DATA_BLOCK "20_TANKS_IP_DATA"   // DB20
TITLE = Tanks Input Data
{ S7_Optimized_Access := 'TRUE' }
AUTHOR : JRS
VERSION : 0.1
// Processed data for code use
   VAR
      RIO_01 : "3T_IP_DATA";   // 1st = FPT, 2nd = 1P, 3rd = 1S
      RIO_02 : "2T_IP_DATA";   // 1st = 2P, 2nd = 2S, 3rd = N/A
      RIO_03 : "2T_IP_DATA";   // 1st = 3P, 2nd = 3S, 3rd = N/A
      RIO_04 : "2T_IP_DATA";   // BWT Level (LT-422)
      RIO_05 : "2T_IP_DATA";   // Raw minimum value from AI card
      RIO_06 : "2T_IP_DATA";   // Raw maximum value from AI card
      RIO_07 : "1T_IP_DATA";   // Normalised real value
   END_VAR
BEGIN
   RIO_02.FIRST_TANK.USD_FLOW_CNFG.ENG_MAX := 500.0;
   RIO_02.FIRST_TANK.MBG_FLOW_CNFG.ENG_MAX := 30.0;
   RIO_02.FIRST_TANK.BWT_PH_CNFG.ENG_MAX := 12.0;
   RIO_02.FIRST_TANK.O2_MONITOR_CNFG.ENG_MAX := 25.0;
   RIO_02.FIRST_TANK.DECK_IG_PRESS_CNFG.ENG_MAX := 10.0;
   RIO_02.FIRST_TANK.TANKS_PRESS_CNFG.ENG_MIN := -200.0;
   RIO_02.FIRST_TANK.TANKS_PRESS_CNFG.ENG_MAX := 200.0;
   RIO_02.FIRST_TANK.BWT_DO_CNFG.ENG_MAX := 20.0;
   RIO_02.FIRST_TANK.BWT_TEMP_CNFG.ENG_MAX := 100.0;
   RIO_02.SECOND_TANK.USD_FLOW_CNFG.ENG_MAX := 500.0;
   RIO_02.SECOND_TANK.MBG_FLOW_CNFG.ENG_MAX := 30.0;
   RIO_02.SECOND_TANK.BWT_PH_CNFG.ENG_MAX := 12.0;
   RIO_02.SECOND_TANK.BWT_DO_CNFG.ENG_MAX := 20.0;
   RIO_02.SECOND_TANK.O2_MONITOR_CNFG.ENG_MAX := 15.0;
   RIO_02.SECOND_TANK.DECK_IG_PRESS_CNFG.ENG_MAX := 25.0;
   RIO_02.SECOND_TANK.TANKS_PRESS_CNFG.ENG_MIN := -200.0;
   RIO_02.SECOND_TANK.TANKS_PRESS_CNFG.ENG_MAX := 200.0;
   RIO_02.SECOND_TANK.BWT_TEMP_CNFG.ENG_MIN := -20.0;
   RIO_02.SECOND_TANK.BWT_TEMP_CNFG.ENG_MAX := 100.0;
   RIO_02.FIRST_TANK.BWT_TEMP_CNFG.ENG_MIN := -20.0;
   RIO_02.FIRST_TANK.BWT_PH_CNFG.ENG_MIN := 2.0;
   RIO_02.SECOND_TANK.BWT_PH_CNFG.ENG_MIN := 2.0;
   RIO_01.FIRST_TANK.O2_MONITOR_CNFG.ENG_MAX := 25.0;   // Engineering units maximum value
   RIO_01.SECOND_TANK.O2_MONITOR_CNFG.ENG_MAX := 25.0;   // Engineering units maximum value
   RIO_01.THIRD_TANK.O2_MONITOR_CNFG.ENG_MAX := 25.0;   // Engineering units maximum value
   RIO_03.FIRST_TANK.O2_MONITOR_CNFG.ENG_MAX := 25.0;   // Engineering units maximum value
   RIO_03.SECOND_TANK.O2_MONITOR_CNFG.ENG_MAX := 25.0;   // Engineering units maximum value
   RIO_04.FIRST_TANK.O2_MONITOR_CNFG.ENG_MAX := 25.0;   // Engineering units maximum value
   RIO_04.SECOND_TANK.O2_MONITOR_CNFG.ENG_MAX := 25.0;   // Engineering units maximum value
   RIO_05.FIRST_TANK.O2_MONITOR_CNFG.ENG_MAX := 25.0;   // Engineering units maximum value
   RIO_05.SECOND_TANK.O2_MONITOR_CNFG.ENG_MAX := 25.0;   // Engineering units maximum value
   RIO_06.FIRST_TANK.O2_MONITOR_CNFG.ENG_MAX := 25.0;   // Engineering units maximum value
   RIO_06.SECOND_TANK.O2_MONITOR_CNFG.ENG_MAX := 25.0;   // Engineering units maximum value
   RIO_07.FIRST_TANK.O2_MONITOR_CNFG.ENG_MAX := 25.0;   // Engineering units maximum value
   RIO_07.FIRST_TANK.BWT_TEMP_CNFG.ENG_MIN := -20.0;   // Engineering units minimum value
   RIO_07.FIRST_TANK.BWT_TEMP_CNFG.ENG_MAX := 100.0;   // Engineering units maximum value
   RIO_07.FIRST_TANK.MBG_FLOW_CNFG.ENG_MAX := 30.0;   // Engineering units maximum value
   RIO_07.FIRST_TANK.USD_FLOW_CNFG.ENG_MAX := 500.0;   // Engineering units maximum value
   RIO_06.FIRST_TANK.BWT_TEMP_CNFG.ENG_MIN := -20.0;   // Engineering units minimum value
   RIO_06.FIRST_TANK.BWT_TEMP_CNFG.ENG_MAX := 100.0;   // Engineering units maximum value
   RIO_06.SECOND_TANK.BWT_TEMP_CNFG.ENG_MIN := -20.0;   // Engineering units minimum value
   RIO_06.SECOND_TANK.BWT_TEMP_CNFG.ENG_MAX := 100.0;   // Engineering units maximum value
   RIO_06.FIRST_TANK.USD_FLOW_CNFG.ENG_MAX := 500.0;   // Engineering units maximum value
   RIO_06.FIRST_TANK.MBG_FLOW_CNFG.ENG_MAX := 30.0;   // Engineering units maximum value
   RIO_06.SECOND_TANK.USD_FLOW_CNFG.ENG_MAX := 500.0;   // Engineering units maximum value
   RIO_06.SECOND_TANK.MBG_FLOW_CNFG.ENG_MAX := 30.0;   // Engineering units maximum value
   RIO_05.FIRST_TANK.BWT_TEMP_CNFG.ENG_MIN := -20.0;   // Engineering units minimum value
   RIO_05.FIRST_TANK.BWT_TEMP_CNFG.ENG_MAX := 100.0;   // Engineering units maximum value
   RIO_05.SECOND_TANK.BWT_TEMP_CNFG.ENG_MIN := -20.0;   // Engineering units minimum value
   RIO_05.SECOND_TANK.BWT_TEMP_CNFG.ENG_MAX := 100.0;   // Engineering units maximum value
   RIO_05.FIRST_TANK.USD_FLOW_CNFG.ENG_MAX := 500.0;   // Engineering units maximum value
   RIO_05.FIRST_TANK.MBG_FLOW_CNFG.ENG_MAX := 30.0;   // Engineering units maximum value
   RIO_05.SECOND_TANK.USD_FLOW_CNFG.ENG_MAX := 500.0;   // Engineering units maximum value
   RIO_05.SECOND_TANK.MBG_FLOW_CNFG.ENG_MAX := 30.0;   // Engineering units maximum value
   RIO_04.FIRST_TANK.USD_FLOW_CNFG.ENG_MAX := 500.0;   // Engineering units maximum value
   RIO_04.FIRST_TANK.MBG_FLOW_CNFG.ENG_MAX := 30.0;   // Engineering units maximum value
   RIO_04.FIRST_TANK.BWT_TEMP_CNFG.ENG_MIN := -20.0;   // Engineering units minimum value
   RIO_04.FIRST_TANK.BWT_TEMP_CNFG.ENG_MAX := 100.0;   // Engineering units maximum value
   RIO_04.SECOND_TANK.USD_FLOW_CNFG.ENG_MAX := 500.0;   // Engineering units maximum value
   RIO_04.SECOND_TANK.MBG_FLOW_CNFG.ENG_MAX := 30.0;   // Engineering units maximum value
   RIO_04.SECOND_TANK.BWT_TEMP_CNFG.ENG_MIN := -20.0;   // Engineering units minimum value
   RIO_04.SECOND_TANK.BWT_TEMP_CNFG.ENG_MAX := 100.0;   // Engineering units maximum value
   RIO_03.FIRST_TANK.USD_FLOW_CNFG.ENG_MAX := 500.0;   // Engineering units maximum value
   RIO_03.FIRST_TANK.MBG_FLOW_CNFG.ENG_MAX := 30.0;   // Engineering units maximum value
   RIO_03.FIRST_TANK.BWT_TEMP_CNFG.ENG_MIN := -20.0;   // Engineering units minimum value
   RIO_03.FIRST_TANK.BWT_TEMP_CNFG.ENG_MAX := 100.0;   // Engineering units maximum value
   RIO_01.FIRST_TANK.USD_FLOW_CNFG.ENG_MAX := 500.0;   // Engineering units maximum value
   RIO_01.FIRST_TANK.MBG_FLOW_CNFG.ENG_MAX := 30.0;   // Engineering units maximum value
   RIO_01.FIRST_TANK.BWT_TEMP_CNFG.ENG_MIN := -20.0;   // Engineering units minimum value
   RIO_01.FIRST_TANK.BWT_TEMP_CNFG.ENG_MAX := 100.0;   // Engineering units maximum value
   RIO_01.SECOND_TANK.USD_FLOW_CNFG.ENG_MAX := 500.0;   // Engineering units maximum value
   RIO_01.SECOND_TANK.MBG_FLOW_CNFG.ENG_MAX := 30.0;   // Engineering units maximum value
   RIO_01.SECOND_TANK.BWT_TEMP_CNFG.ENG_MIN := -20.0;   // Engineering units minimum value
   RIO_01.SECOND_TANK.BWT_TEMP_CNFG.ENG_MAX := 100.0;   // Engineering units maximum value
   RIO_01.THIRD_TANK.USD_FLOW_CNFG.ENG_MAX := 500.0;   // Engineering units maximum value
   RIO_01.THIRD_TANK.MBG_FLOW_CNFG.ENG_MAX := 30.0;   // Engineering units maximum value
   RIO_01.THIRD_TANK.BWT_TEMP_CNFG.ENG_MIN := -20.0;   // Engineering units minimum value
   RIO_01.THIRD_TANK.BWT_TEMP_CNFG.ENG_MAX := 100.0;   // Engineering units maximum value
   RIO_03.SECOND_TANK.USD_FLOW_CNFG.ENG_MAX := 500.0;   // Engineering units maximum value
   RIO_03.SECOND_TANK.MBG_FLOW_CNFG.ENG_MAX := 30.0;   // Engineering units maximum value
   // RIO_02.FIRST_TANK.USD_FLOW_CNFG : IW160 - USD Flow (FIT-418) - Tank #1
   // RIO_02.FIRST_TANK.MBG_FLOW_CNFG : IW162 - MBG Flow (FIT-420) - Tank #1
   // RIO_02.FIRST_TANK.BWT_LEVEL_CNFG : BWT Level (LT-422)
   // RIO_02.FIRST_TANK.BWT_PH_CNFG : BWT Ph (426)
   // RIO_02.FIRST_TANK.BWT_TEMP_CNFG : BWT Temperature (426)
   // RIO_02.FIRST_TANK.BWT_DO_CNFG : BWT DO (428)
   // RIO_02.FIRST_TANK.O2_MONITOR_CNFG : O2 Monitor (600-Tx-433)
   // RIO_02.FIRST_TANK.DECK_IG_PRESS_CNFG : Deck Main IG Pressure (PT-415)
   // RIO_02.FIRST_TANK.TANKS_PRESS_CNFG : Tank Group Pressure (PT-424)
   // RIO_02.SECOND_TANK.USD_FLOW_CNFG : IW160 - USD Flow (FIT-417) - Tank #1
   // RIO_02.SECOND_TANK.MBG_FLOW_CNFG : IW162 - MBG Flow (FIT-419) - Tank #1
   // RIO_02.SECOND_TANK.BWT_LEVEL_CNFG : BWT Level (LT-422)
   // RIO_02.SECOND_TANK.BWT_PH_CNFG : BWT Ph (426)
   // RIO_02.SECOND_TANK.BWT_TEMP_CNFG : BWT Temperature (426)
   // RIO_02.SECOND_TANK.BWT_DO_CNFG : BWT DO (428)
   // RIO_02.SECOND_TANK.SPARE_AI_1_CNFG : Input processing configuration data
   // RIO_02.SECOND_TANK.SPARE_AI_2_CNFG : Input processing configuration data
   // RIO_02.SECOND_TANK.SPARE_AI_3_CNFG : Input processing configuration data
   // RIO_02.SECOND_TANK.O2_MONITOR_CNFG : O2 Monitor (600-Tx-433)
   // RIO_02.SECOND_TANK.DECK_IG_PRESS_CNFG : Deck Main IG Pressure (PT-415)
   // RIO_02.SECOND_TANK.TANKS_PRESS_CNFG : Tank Group Pressure (PT-424)
   // RIO_02.SECOND_TANK.MBG_FLOW : FIT-419
   // RIO_02.SECOND_TANK.USD_FLOW : FIT-417
   // RIO_01.FIRST_TANK.O2_MONITOR : Space monitor, 600-Tx-433
   // RIO_01.FIRST_TANK.DECK_IG_PRESS : Deck main IG pressure, PT-415
   // RIO_01.FIRST_TANK.TANKS_PRESS : Tank group pressure, PT-424
   // RIO_01.FIRST_TANK.TANKS_PRESS_HIHI : Tank group pressure, PS-436
   // RIO_01.FIRST_TANK.TANK_GROUP_SPARE_DI_2 : Spare input
   // RIO_01.FIRST_TANK.TANK_GROUP_SPARE_DI_3 : Spare input
   // RIO_01.FIRST_TANK.TANK_GROUP_SPARE_DI_4 : Spare input
   // RIO_01.FIRST_TANK.TANK_GROUP_SPARE_DI_5 : Spare input
   // RIO_01.FIRST_TANK.TANK_GROUP_SPARE_DI_6 : Spare input
   // RIO_01.FIRST_TANK.TANK_GROUP_SPARE_DI_7 : Spare input
   // RIO_01.FIRST_TANK.GTT_ISOL_VALVE_OPEN : Gas to tank isolation valve feedback, CV-422
   // RIO_01.FIRST_TANK.GTT_ISOL_VALVE_CLSD : Gas to tank isolation valve feedback, CV-422
   // RIO_01.FIRST_TANK.TANK_VENT_A_OPEN : Tank vent valve feedback, CV-441-A
   // RIO_01.FIRST_TANK.TANK_VENT_A_CLSD : Tank vent valve feedback, CV-441-A
   // RIO_01.FIRST_TANK.TANK_VENT_B_OPEN : Tank vent valve feedback, CV-441-B
   // RIO_01.FIRST_TANK.TANK_VENT_B_CLSD : Tank vent valve feedback, CV-441-B
   // RIO_01.FIRST_TANK.BWT_LEVEL_HIHI : Tank water level, LS-425
   // RIO_01.FIRST_TANK.TANK_ALARM : Spare input
   // RIO_01.FIRST_TANK.SPARE_DI_7 : Spare input
   // RIO_01.FIRST_TANK.USD_FLOW : FIT-418
   // RIO_01.FIRST_TANK.MBG_FLOW : FIT-420
   // RIO_01.FIRST_TANK.BWT_LEVEL : LT-422
   // RIO_01.FIRST_TANK.BWT_PH : Ph 426
   // RIO_01.FIRST_TANK.BWT_TEMP : Temperature 426
   // RIO_01.FIRST_TANK.BWT_DO : Disolved oxygen 428
   // RIO_01.FIRST_TANK.SPARE_AI_1 : Spare input
   // RIO_01.FIRST_TANK.SPARE_AI_2 : Spare input
   // RIO_01.FIRST_TANK.SPARE_AI_3 : Spare input
   // RIO_01.FIRST_TANK.USD_FLOW_CNFG : IW160 - USD Flow (FIT-418) - Tank #1
   // RIO_01.FIRST_TANK.USD_FLOW_CNFG.RAW_MIN : Raw minimum value from AI card
   // RIO_01.FIRST_TANK.USD_FLOW_CNFG.RAW_MAX : Raw maximum value from AI card
   // RIO_01.FIRST_TANK.USD_FLOW_CNFG.NORM : Normalised real value
   // RIO_01.FIRST_TANK.USD_FLOW_CNFG.ENG_MIN : Engineering units minimum value
   // RIO_01.FIRST_TANK.MBG_FLOW_CNFG : IW162 - MBG Flow (FIT-420) - Tank #1
   // RIO_01.FIRST_TANK.MBG_FLOW_CNFG.RAW_MIN : Raw minimum value from AI card
   // RIO_01.FIRST_TANK.MBG_FLOW_CNFG.RAW_MAX : Raw maximum value from AI card
   // RIO_01.FIRST_TANK.MBG_FLOW_CNFG.NORM : Normalised real value
   // RIO_01.FIRST_TANK.MBG_FLOW_CNFG.ENG_MIN : Engineering units minimum value
   // RIO_01.FIRST_TANK.BWT_LEVEL_CNFG : BWT Level (LT-422)
   // RIO_01.FIRST_TANK.BWT_LEVEL_CNFG.RAW_MIN : Raw minimum value from AI card
   // RIO_01.FIRST_TANK.BWT_LEVEL_CNFG.RAW_MAX : Raw maximum value from AI card
   // RIO_01.FIRST_TANK.BWT_LEVEL_CNFG.NORM : Normalised real value
   // RIO_01.FIRST_TANK.BWT_LEVEL_CNFG.ENG_MIN : Engineering units minimum value
   // RIO_01.FIRST_TANK.BWT_LEVEL_CNFG.ENG_MAX : Engineering units maximum value
   // RIO_01.FIRST_TANK.BWT_PH_CNFG : BWT Ph (426)
   // RIO_01.FIRST_TANK.BWT_PH_CNFG.RAW_MIN : Raw minimum value from AI card
   // RIO_01.FIRST_TANK.BWT_PH_CNFG.RAW_MAX : Raw maximum value from AI card
   // RIO_01.FIRST_TANK.BWT_PH_CNFG.NORM : Normalised real value
   // RIO_01.FIRST_TANK.BWT_PH_CNFG.ENG_MIN : Engineering units minimum value
   // RIO_01.FIRST_TANK.BWT_PH_CNFG.ENG_MAX : Engineering units maximum value
   // RIO_01.FIRST_TANK.BWT_TEMP_CNFG : BWT Temperature (426)
   // RIO_01.FIRST_TANK.BWT_TEMP_CNFG.RAW_MIN : Raw minimum value from AI card
   // RIO_01.FIRST_TANK.BWT_TEMP_CNFG.RAW_MAX : Raw maximum value from AI card
   // RIO_01.FIRST_TANK.BWT_TEMP_CNFG.NORM : Normalised real value
   // RIO_01.FIRST_TANK.BWT_DO_CNFG : BWT DO (428)
   // RIO_01.FIRST_TANK.BWT_DO_CNFG.RAW_MIN : Raw minimum value from AI card
   // RIO_01.FIRST_TANK.BWT_DO_CNFG.RAW_MAX : Raw maximum value from AI card
   // RIO_01.FIRST_TANK.BWT_DO_CNFG.NORM : Normalised real value
   // RIO_01.FIRST_TANK.BWT_DO_CNFG.ENG_MIN : Engineering units minimum value
   // RIO_01.FIRST_TANK.BWT_DO_CNFG.ENG_MAX : Engineering units maximum value
   // RIO_01.FIRST_TANK.SPARE_AI_1_CNFG : Input processing configuration data
   // RIO_01.FIRST_TANK.SPARE_AI_1_CNFG.RAW_MIN : Raw minimum value from AI card
   // RIO_01.FIRST_TANK.SPARE_AI_1_CNFG.RAW_MAX : Raw maximum value from AI card
   // RIO_01.FIRST_TANK.SPARE_AI_1_CNFG.NORM : Normalised real value
   // RIO_01.FIRST_TANK.SPARE_AI_1_CNFG.ENG_MIN : Engineering units minimum value
   // RIO_01.FIRST_TANK.SPARE_AI_1_CNFG.ENG_MAX : Engineering units maximum value
   // RIO_01.FIRST_TANK.SPARE_AI_2_CNFG : Input processing configuration data
   // RIO_01.FIRST_TANK.SPARE_AI_2_CNFG.RAW_MIN : Raw minimum value from AI card
   // RIO_01.FIRST_TANK.SPARE_AI_2_CNFG.RAW_MAX : Raw maximum value from AI card
   // RIO_01.FIRST_TANK.SPARE_AI_2_CNFG.NORM : Normalised real value
   // RIO_01.FIRST_TANK.SPARE_AI_2_CNFG.ENG_MIN : Engineering units minimum value
   // RIO_01.FIRST_TANK.SPARE_AI_2_CNFG.ENG_MAX : Engineering units maximum value
   // RIO_01.FIRST_TANK.SPARE_AI_3_CNFG : Input processing configuration data
   // RIO_01.FIRST_TANK.SPARE_AI_3_CNFG.RAW_MIN : Raw minimum value from AI card
   // RIO_01.FIRST_TANK.SPARE_AI_3_CNFG.RAW_MAX : Raw maximum value from AI card
   // RIO_01.FIRST_TANK.SPARE_AI_3_CNFG.NORM : Normalised real value
   // RIO_01.FIRST_TANK.SPARE_AI_3_CNFG.ENG_MIN : Engineering units minimum value
   // RIO_01.FIRST_TANK.SPARE_AI_3_CNFG.ENG_MAX : Engineering units maximum value
   // RIO_01.FIRST_TANK.O2_MONITOR_CNFG : O2 Monitor (600-Tx-433)
   // RIO_01.FIRST_TANK.O2_MONITOR_CNFG.RAW_MIN : Raw minimum value from AI card
   // RIO_01.FIRST_TANK.O2_MONITOR_CNFG.RAW_MAX : Raw maximum value from AI card
   // RIO_01.FIRST_TANK.O2_MONITOR_CNFG.NORM : Normalised real value
   // RIO_01.FIRST_TANK.O2_MONITOR_CNFG.ENG_MIN : Engineering units minimum value
   // RIO_01.FIRST_TANK.DECK_IG_PRESS_CNFG : Deck Main IG Pressure (PT-415)
   // RIO_01.FIRST_TANK.DECK_IG_PRESS_CNFG.RAW_MIN : Raw minimum value from AI card
   // RIO_01.FIRST_TANK.DECK_IG_PRESS_CNFG.RAW_MAX : Raw maximum value from AI card
   // RIO_01.FIRST_TANK.DECK_IG_PRESS_CNFG.NORM : Normalised real value
   // RIO_01.FIRST_TANK.DECK_IG_PRESS_CNFG.ENG_MIN : Engineering units minimum value
   // RIO_01.FIRST_TANK.DECK_IG_PRESS_CNFG.ENG_MAX : Engineering units maximum value
   // RIO_01.FIRST_TANK.TANKS_PRESS_CNFG : Tank Group Pressure (PT-424)
   // RIO_01.FIRST_TANK.TANKS_PRESS_CNFG.RAW_MIN : Raw minimum value from AI card
   // RIO_01.FIRST_TANK.TANKS_PRESS_CNFG.RAW_MAX : Raw maximum value from AI card
   // RIO_01.FIRST_TANK.TANKS_PRESS_CNFG.NORM : Normalised real value
   // RIO_01.FIRST_TANK.TANKS_PRESS_CNFG.ENG_MIN : Engineering units minimum value
   // RIO_01.FIRST_TANK.TANKS_PRESS_CNFG.ENG_MAX : Engineering units maximum value
   // RIO_01.THIRD_TANK.O2_MONITOR : Space monitor, 600-Tx-433
   // RIO_01.THIRD_TANK.DECK_IG_PRESS : Deck main IG pressure, PT-415
   // RIO_01.THIRD_TANK.TANKS_PRESS : Tank group pressure, PT-424
   // RIO_01.THIRD_TANK.TANKS_PRESS_HIHI : Tank group pressure, PS-436
   // RIO_01.THIRD_TANK.TANK_GROUP_SPARE_DI_2 : Spare input
   // RIO_01.THIRD_TANK.TANK_GROUP_SPARE_DI_3 : Spare input
   // RIO_01.THIRD_TANK.TANK_GROUP_SPARE_DI_4 : Spare input
   // RIO_01.THIRD_TANK.TANK_GROUP_SPARE_DI_5 : Spare input
   // RIO_01.THIRD_TANK.TANK_GROUP_SPARE_DI_6 : Spare input
   // RIO_01.THIRD_TANK.TANK_GROUP_SPARE_DI_7 : Spare input
   // RIO_01.THIRD_TANK.GTT_ISOL_VALVE_OPEN : Gas to tank isolation valve feedback, CV-422
   // RIO_01.THIRD_TANK.GTT_ISOL_VALVE_CLSD : Gas to tank isolation valve feedback, CV-422
   // RIO_01.THIRD_TANK.TANK_VENT_A_OPEN : Tank vent valve feedback, CV-441-A
   // RIO_01.THIRD_TANK.TANK_VENT_A_CLSD : Tank vent valve feedback, CV-441-A
   // RIO_01.THIRD_TANK.TANK_VENT_B_OPEN : Tank vent valve feedback, CV-441-B
   // RIO_01.THIRD_TANK.TANK_VENT_B_CLSD : Tank vent valve feedback, CV-441-B
   // RIO_01.THIRD_TANK.BWT_LEVEL_HIHI : Tank water level, LS-425
   // RIO_01.THIRD_TANK.TANK_ALARM : Spare input
   // RIO_01.THIRD_TANK.SPARE_DI_7 : Spare input
   // RIO_01.THIRD_TANK.USD_FLOW : FIT-417
   // RIO_01.THIRD_TANK.MBG_FLOW : FIT-419
   // RIO_01.THIRD_TANK.BWT_LEVEL : LT-422
   // RIO_01.THIRD_TANK.BWT_PH : Ph 426
   // RIO_01.THIRD_TANK.BWT_TEMP : Temperature 426
   // RIO_01.THIRD_TANK.BWT_DO : Disolved oxygen 428
   // RIO_01.THIRD_TANK.SPARE_AI_1 : Spare input
   // RIO_01.THIRD_TANK.SPARE_AI_2 : Spare input
   // RIO_01.THIRD_TANK.SPARE_AI_3 : Spare input
   // RIO_01.THIRD_TANK.USD_FLOW_CNFG : IW160 - USD Flow (FIT-417) - Tank #1
   // RIO_01.THIRD_TANK.USD_FLOW_CNFG.RAW_MIN : Raw minimum value from AI card
   // RIO_01.THIRD_TANK.USD_FLOW_CNFG.RAW_MAX : Raw maximum value from AI card
   // RIO_01.THIRD_TANK.USD_FLOW_CNFG.NORM : Normalised real value
   // RIO_01.THIRD_TANK.USD_FLOW_CNFG.ENG_MIN : Engineering units minimum value
   // RIO_01.THIRD_TANK.MBG_FLOW_CNFG : IW162 - MBG Flow (FIT-420) - Tank #1
   // RIO_01.THIRD_TANK.MBG_FLOW_CNFG.RAW_MIN : Raw minimum value from AI card
   // RIO_01.THIRD_TANK.MBG_FLOW_CNFG.RAW_MAX : Raw maximum value from AI card
   // RIO_01.THIRD_TANK.MBG_FLOW_CNFG.NORM : Normalised real value
   // RIO_01.THIRD_TANK.MBG_FLOW_CNFG.ENG_MIN : Engineering units minimum value
   // RIO_01.THIRD_TANK.BWT_LEVEL_CNFG : BWT Level (LT-422)
   // RIO_01.THIRD_TANK.BWT_LEVEL_CNFG.RAW_MIN : Raw minimum value from AI card
   // RIO_01.THIRD_TANK.BWT_LEVEL_CNFG.RAW_MAX : Raw maximum value from AI card
   // RIO_01.THIRD_TANK.BWT_LEVEL_CNFG.NORM : Normalised real value
   // RIO_01.THIRD_TANK.BWT_LEVEL_CNFG.ENG_MIN : Engineering units minimum value
   // RIO_01.THIRD_TANK.BWT_LEVEL_CNFG.ENG_MAX : Engineering units maximum value
   // RIO_01.THIRD_TANK.BWT_PH_CNFG : BWT Ph (426)
   // RIO_01.THIRD_TANK.BWT_PH_CNFG.RAW_MIN : Raw minimum value from AI card
   // RIO_01.THIRD_TANK.BWT_PH_CNFG.RAW_MAX : Raw maximum value from AI card
   // RIO_01.THIRD_TANK.BWT_PH_CNFG.NORM : Normalised real value
   // RIO_01.THIRD_TANK.BWT_PH_CNFG.ENG_MIN : Engineering units minimum value
   // RIO_01.THIRD_TANK.BWT_PH_CNFG.ENG_MAX : Engineering units maximum value
   // RIO_01.THIRD_TANK.BWT_TEMP_CNFG : BWT Temperature (426)
   // RIO_01.THIRD_TANK.BWT_TEMP_CNFG.RAW_MIN : Raw minimum value from AI card
   // RIO_01.THIRD_TANK.BWT_TEMP_CNFG.RAW_MAX : Raw maximum value from AI card
   // RIO_01.THIRD_TANK.BWT_TEMP_CNFG.NORM : Normalised real value
   // RIO_01.THIRD_TANK.BWT_DO_CNFG : BWT DO (428)
   // RIO_01.THIRD_TANK.BWT_DO_CNFG.RAW_MIN : Raw minimum value from AI card
   // RIO_01.THIRD_TANK.BWT_DO_CNFG.RAW_MAX : Raw maximum value from AI card
   // RIO_01.THIRD_TANK.BWT_DO_CNFG.NORM : Normalised real value
   // RIO_01.THIRD_TANK.BWT_DO_CNFG.ENG_MIN : Engineering units minimum value
   // RIO_01.THIRD_TANK.BWT_DO_CNFG.ENG_MAX : Engineering units maximum value
   // RIO_01.THIRD_TANK.SPARE_AI_1_CNFG : Input processing configuration data
   // RIO_01.THIRD_TANK.SPARE_AI_1_CNFG.RAW_MIN : Raw minimum value from AI card
   // RIO_01.THIRD_TANK.SPARE_AI_1_CNFG.RAW_MAX : Raw maximum value from AI card
   // RIO_01.THIRD_TANK.SPARE_AI_1_CNFG.NORM : Normalised real value
   // RIO_01.THIRD_TANK.SPARE_AI_1_CNFG.ENG_MIN : Engineering units minimum value
   // RIO_01.THIRD_TANK.SPARE_AI_1_CNFG.ENG_MAX : Engineering units maximum value
   // RIO_01.THIRD_TANK.SPARE_AI_2_CNFG : Input processing configuration data
   // RIO_01.THIRD_TANK.SPARE_AI_2_CNFG.RAW_MIN : Raw minimum value from AI card
   // RIO_01.THIRD_TANK.SPARE_AI_2_CNFG.RAW_MAX : Raw maximum value from AI card
   // RIO_01.THIRD_TANK.SPARE_AI_2_CNFG.NORM : Normalised real value
   // RIO_01.THIRD_TANK.SPARE_AI_2_CNFG.ENG_MIN : Engineering units minimum value
   // RIO_01.THIRD_TANK.SPARE_AI_2_CNFG.ENG_MAX : Engineering units maximum value
   // RIO_01.THIRD_TANK.SPARE_AI_3_CNFG : Input processing configuration data
   // RIO_01.THIRD_TANK.SPARE_AI_3_CNFG.RAW_MIN : Raw minimum value from AI card
   // RIO_01.THIRD_TANK.SPARE_AI_3_CNFG.RAW_MAX : Raw maximum value from AI card
   // RIO_01.THIRD_TANK.SPARE_AI_3_CNFG.NORM : Normalised real value
   // RIO_01.THIRD_TANK.SPARE_AI_3_CNFG.ENG_MIN : Engineering units minimum value
   // RIO_01.THIRD_TANK.SPARE_AI_3_CNFG.ENG_MAX : Engineering units maximum value
   // RIO_01.THIRD_TANK.O2_MONITOR_CNFG : O2 Monitor (600-Tx-433)
   // RIO_01.THIRD_TANK.O2_MONITOR_CNFG.RAW_MIN : Raw minimum value from AI card
   // RIO_01.THIRD_TANK.O2_MONITOR_CNFG.RAW_MAX : Raw maximum value from AI card
   // RIO_01.THIRD_TANK.O2_MONITOR_CNFG.NORM : Normalised real value
   // RIO_01.THIRD_TANK.O2_MONITOR_CNFG.ENG_MIN : Engineering units minimum value
   // RIO_01.THIRD_TANK.DECK_IG_PRESS_CNFG : Deck Main IG Pressure (PT-415)
   // RIO_01.THIRD_TANK.DECK_IG_PRESS_CNFG.RAW_MIN : Raw minimum value from AI card
   // RIO_01.THIRD_TANK.DECK_IG_PRESS_CNFG.RAW_MAX : Raw maximum value from AI card
   // RIO_01.THIRD_TANK.DECK_IG_PRESS_CNFG.NORM : Normalised real value
   // RIO_01.THIRD_TANK.DECK_IG_PRESS_CNFG.ENG_MIN : Engineering units minimum value
   // RIO_01.THIRD_TANK.DECK_IG_PRESS_CNFG.ENG_MAX : Engineering units maximum value
   // RIO_01.THIRD_TANK.TANKS_PRESS_CNFG : Tank Group Pressure (PT-424)
   // RIO_01.THIRD_TANK.TANKS_PRESS_CNFG.RAW_MIN : Raw minimum value from AI card
   // RIO_01.THIRD_TANK.TANKS_PRESS_CNFG.RAW_MAX : Raw maximum value from AI card
   // RIO_01.THIRD_TANK.TANKS_PRESS_CNFG.NORM : Normalised real value
   // RIO_01.THIRD_TANK.TANKS_PRESS_CNFG.ENG_MIN : Engineering units minimum value
   // RIO_01.THIRD_TANK.TANKS_PRESS_CNFG.ENG_MAX : Engineering units maximum value
   // RIO_03.SECOND_TANK.O2_MONITOR : Space monitor, 600-Tx-433
   // RIO_03.SECOND_TANK.DECK_IG_PRESS : Deck main IG pressure, PT-415
   // RIO_03.SECOND_TANK.TANKS_PRESS : Tank group pressure, PT-424
   // RIO_03.SECOND_TANK.TANKS_PRESS_HIHI : Tank group pressure, PS-436
   // RIO_03.SECOND_TANK.TANK_GROUP_SPARE_DI_2 : Spare input
   // RIO_03.SECOND_TANK.TANK_GROUP_SPARE_DI_3 : Spare input
   // RIO_03.SECOND_TANK.TANK_GROUP_SPARE_DI_4 : Spare input
   // RIO_03.SECOND_TANK.TANK_GROUP_SPARE_DI_5 : Spare input
   // RIO_03.SECOND_TANK.TANK_GROUP_SPARE_DI_6 : Spare input
   // RIO_03.SECOND_TANK.TANK_GROUP_SPARE_DI_7 : Spare input
   // RIO_03.SECOND_TANK.GTT_ISOL_VALVE_OPEN : Gas to tank isolation valve feedback, CV-422
   // RIO_03.SECOND_TANK.GTT_ISOL_VALVE_CLSD : Gas to tank isolation valve feedback, CV-422
   // RIO_03.SECOND_TANK.TANK_VENT_A_OPEN : Tank vent valve feedback, CV-441-A
   // RIO_03.SECOND_TANK.TANK_VENT_A_CLSD : Tank vent valve feedback, CV-441-A
   // RIO_03.SECOND_TANK.TANK_VENT_B_OPEN : Tank vent valve feedback, CV-441-B
   // RIO_03.SECOND_TANK.TANK_VENT_B_CLSD : Tank vent valve feedback, CV-441-B
   // RIO_03.SECOND_TANK.BWT_LEVEL_HIHI : Tank water level, LS-425
   // RIO_03.SECOND_TANK.TANK_ALARM : Spare input
   // RIO_03.SECOND_TANK.SPARE_DI_7 : Spare input
   // RIO_03.SECOND_TANK.USD_FLOW : FIT-417
   // RIO_03.SECOND_TANK.MBG_FLOW : FIT-419
   // RIO_03.SECOND_TANK.BWT_LEVEL : LT-422
   // RIO_03.SECOND_TANK.BWT_PH : Ph 426
   // RIO_03.SECOND_TANK.BWT_TEMP : Temperature 426
   // RIO_03.SECOND_TANK.BWT_DO : Disolved oxygen 428
   // RIO_03.SECOND_TANK.SPARE_AI_1 : Spare input
   // RIO_03.SECOND_TANK.SPARE_AI_2 : Spare input
   // RIO_03.SECOND_TANK.SPARE_AI_3 : Spare input
   // RIO_03.SECOND_TANK.USD_FLOW_CNFG : IW160 - USD Flow (FIT-417) - Tank #1
   // RIO_03.SECOND_TANK.MBG_FLOW_CNFG : IW162 - MBG Flow (FIT-420) - Tank #1
   // RIO_03.SECOND_TANK.BWT_LEVEL_CNFG : BWT Level (LT-422)
   // RIO_03.SECOND_TANK.BWT_PH_CNFG : BWT Ph (426)
   // RIO_03.SECOND_TANK.BWT_TEMP_CNFG : BWT Temperature (426)
   // RIO_03.SECOND_TANK.BWT_DO_CNFG : BWT DO (428)
   // RIO_03.SECOND_TANK.SPARE_AI_1_CNFG : Input processing configuration data
   // RIO_03.SECOND_TANK.SPARE_AI_2_CNFG : Input processing configuration data
   // RIO_03.SECOND_TANK.SPARE_AI_3_CNFG : Input processing configuration data
   // RIO_03.SECOND_TANK.O2_MONITOR_CNFG : O2 Monitor (600-Tx-433)
   // RIO_03.SECOND_TANK.DECK_IG_PRESS_CNFG : Deck Main IG Pressure (PT-415)
   // RIO_03.SECOND_TANK.TANKS_PRESS_CNFG : Tank Group Pressure (PT-424)
   // RIO_03.FIRST_TANK.O2_MONITOR : Space monitor, 600-Tx-433
   // RIO_03.FIRST_TANK.DECK_IG_PRESS : Deck main IG pressure, PT-415
   // RIO_03.FIRST_TANK.TANKS_PRESS : Tank group pressure, PT-424
   // RIO_03.FIRST_TANK.TANKS_PRESS_HIHI : Tank group pressure, PS-436
   // RIO_03.FIRST_TANK.TANK_GROUP_SPARE_DI_2 : Spare input
   // RIO_03.FIRST_TANK.TANK_GROUP_SPARE_DI_3 : Spare input
   // RIO_03.FIRST_TANK.TANK_GROUP_SPARE_DI_4 : Spare input
   // RIO_03.FIRST_TANK.TANK_GROUP_SPARE_DI_5 : Spare input
   // RIO_03.FIRST_TANK.TANK_GROUP_SPARE_DI_6 : Spare input
   // RIO_03.FIRST_TANK.TANK_GROUP_SPARE_DI_7 : Spare input
   // RIO_03.FIRST_TANK.GTT_ISOL_VALVE_OPEN : Gas to tank isolation valve feedback, CV-422
   // RIO_03.FIRST_TANK.GTT_ISOL_VALVE_CLSD : Gas to tank isolation valve feedback, CV-422
   // RIO_03.FIRST_TANK.TANK_VENT_A_OPEN : Tank vent valve feedback, CV-441-A
   // RIO_03.FIRST_TANK.TANK_VENT_A_CLSD : Tank vent valve feedback, CV-441-A
   // RIO_03.FIRST_TANK.TANK_VENT_B_OPEN : Tank vent valve feedback, CV-441-B
   // RIO_03.FIRST_TANK.TANK_VENT_B_CLSD : Tank vent valve feedback, CV-441-B
   // RIO_03.FIRST_TANK.BWT_LEVEL_HIHI : Tank water level, LS-425
   // RIO_03.FIRST_TANK.TANK_ALARM : Spare input
   // RIO_03.FIRST_TANK.SPARE_DI_7 : Spare input
   // RIO_03.FIRST_TANK.USD_FLOW : FIT-418
   // RIO_03.FIRST_TANK.MBG_FLOW : FIT-420
   // RIO_03.FIRST_TANK.BWT_LEVEL : LT-422
   // RIO_03.FIRST_TANK.BWT_PH : Ph 426
   // RIO_03.FIRST_TANK.BWT_TEMP : Temperature 426
   // RIO_03.FIRST_TANK.BWT_DO : Disolved oxygen 428
   // RIO_03.FIRST_TANK.SPARE_AI_1 : Spare input
   // RIO_03.FIRST_TANK.SPARE_AI_2 : Spare input
   // RIO_03.FIRST_TANK.SPARE_AI_3 : Spare input
   // RIO_03.FIRST_TANK.USD_FLOW_CNFG : IW160 - USD Flow (FIT-418) - Tank #1
   // RIO_03.FIRST_TANK.USD_FLOW_CNFG.RAW_MIN : Raw minimum value from AI card
   // RIO_03.FIRST_TANK.USD_FLOW_CNFG.RAW_MAX : Raw maximum value from AI card
   // RIO_03.FIRST_TANK.USD_FLOW_CNFG.NORM : Normalised real value
   // RIO_03.FIRST_TANK.USD_FLOW_CNFG.ENG_MIN : Engineering units minimum value
   // RIO_03.FIRST_TANK.MBG_FLOW_CNFG : IW162 - MBG Flow (FIT-420) - Tank #1
   // RIO_03.FIRST_TANK.MBG_FLOW_CNFG.RAW_MIN : Raw minimum value from AI card
   // RIO_03.FIRST_TANK.MBG_FLOW_CNFG.RAW_MAX : Raw maximum value from AI card
   // RIO_03.FIRST_TANK.MBG_FLOW_CNFG.NORM : Normalised real value
   // RIO_03.FIRST_TANK.MBG_FLOW_CNFG.ENG_MIN : Engineering units minimum value
   // RIO_03.FIRST_TANK.BWT_LEVEL_CNFG : BWT Level (LT-422)
   // RIO_03.FIRST_TANK.BWT_LEVEL_CNFG.RAW_MIN : Raw minimum value from AI card
   // RIO_03.FIRST_TANK.BWT_LEVEL_CNFG.RAW_MAX : Raw maximum value from AI card
   // RIO_03.FIRST_TANK.BWT_LEVEL_CNFG.NORM : Normalised real value
   // RIO_03.FIRST_TANK.BWT_LEVEL_CNFG.ENG_MIN : Engineering units minimum value
   // RIO_03.FIRST_TANK.BWT_LEVEL_CNFG.ENG_MAX : Engineering units maximum value
   // RIO_03.FIRST_TANK.BWT_PH_CNFG : BWT Ph (426)
   // RIO_03.FIRST_TANK.BWT_PH_CNFG.RAW_MIN : Raw minimum value from AI card
   // RIO_03.FIRST_TANK.BWT_PH_CNFG.RAW_MAX : Raw maximum value from AI card
   // RIO_03.FIRST_TANK.BWT_PH_CNFG.NORM : Normalised real value
   // RIO_03.FIRST_TANK.BWT_PH_CNFG.ENG_MIN : Engineering units minimum value
   // RIO_03.FIRST_TANK.BWT_PH_CNFG.ENG_MAX : Engineering units maximum value
   // RIO_03.FIRST_TANK.BWT_TEMP_CNFG : BWT Temperature (426)
   // RIO_03.FIRST_TANK.BWT_TEMP_CNFG.RAW_MIN : Raw minimum value from AI card
   // RIO_03.FIRST_TANK.BWT_TEMP_CNFG.RAW_MAX : Raw maximum value from AI card
   // RIO_03.FIRST_TANK.BWT_TEMP_CNFG.NORM : Normalised real value
   // RIO_03.FIRST_TANK.BWT_DO_CNFG : BWT DO (428)
   // RIO_03.FIRST_TANK.BWT_DO_CNFG.RAW_MIN : Raw minimum value from AI card
   // RIO_03.FIRST_TANK.BWT_DO_CNFG.RAW_MAX : Raw maximum value from AI card
   // RIO_03.FIRST_TANK.BWT_DO_CNFG.NORM : Normalised real value
   // RIO_03.FIRST_TANK.BWT_DO_CNFG.ENG_MIN : Engineering units minimum value
   // RIO_03.FIRST_TANK.BWT_DO_CNFG.ENG_MAX : Engineering units maximum value
   // RIO_03.FIRST_TANK.SPARE_AI_1_CNFG : Input processing configuration data
   // RIO_03.FIRST_TANK.SPARE_AI_1_CNFG.RAW_MIN : Raw minimum value from AI card
   // RIO_03.FIRST_TANK.SPARE_AI_1_CNFG.RAW_MAX : Raw maximum value from AI card
   // RIO_03.FIRST_TANK.SPARE_AI_1_CNFG.NORM : Normalised real value
   // RIO_03.FIRST_TANK.SPARE_AI_1_CNFG.ENG_MIN : Engineering units minimum value
   // RIO_03.FIRST_TANK.SPARE_AI_1_CNFG.ENG_MAX : Engineering units maximum value
   // RIO_03.FIRST_TANK.SPARE_AI_2_CNFG : Input processing configuration data
   // RIO_03.FIRST_TANK.SPARE_AI_2_CNFG.RAW_MIN : Raw minimum value from AI card
   // RIO_03.FIRST_TANK.SPARE_AI_2_CNFG.RAW_MAX : Raw maximum value from AI card
   // RIO_03.FIRST_TANK.SPARE_AI_2_CNFG.NORM : Normalised real value
   // RIO_03.FIRST_TANK.SPARE_AI_2_CNFG.ENG_MIN : Engineering units minimum value
   // RIO_03.FIRST_TANK.SPARE_AI_2_CNFG.ENG_MAX : Engineering units maximum value
   // RIO_03.FIRST_TANK.SPARE_AI_3_CNFG : Input processing configuration data
   // RIO_03.FIRST_TANK.SPARE_AI_3_CNFG.RAW_MIN : Raw minimum value from AI card
   // RIO_03.FIRST_TANK.SPARE_AI_3_CNFG.RAW_MAX : Raw maximum value from AI card
   // RIO_03.FIRST_TANK.SPARE_AI_3_CNFG.NORM : Normalised real value
   // RIO_03.FIRST_TANK.SPARE_AI_3_CNFG.ENG_MIN : Engineering units minimum value
   // RIO_03.FIRST_TANK.SPARE_AI_3_CNFG.ENG_MAX : Engineering units maximum value
   // RIO_03.FIRST_TANK.O2_MONITOR_CNFG : O2 Monitor (600-Tx-433)
   // RIO_03.FIRST_TANK.O2_MONITOR_CNFG.RAW_MIN : Raw minimum value from AI card
   // RIO_03.FIRST_TANK.O2_MONITOR_CNFG.RAW_MAX : Raw maximum value from AI card
   // RIO_03.FIRST_TANK.O2_MONITOR_CNFG.NORM : Normalised real value
   // RIO_03.FIRST_TANK.O2_MONITOR_CNFG.ENG_MIN : Engineering units minimum value
   // RIO_03.FIRST_TANK.DECK_IG_PRESS_CNFG : Deck Main IG Pressure (PT-415)
   // RIO_03.FIRST_TANK.DECK_IG_PRESS_CNFG.RAW_MIN : Raw minimum value from AI card
   // RIO_03.FIRST_TANK.DECK_IG_PRESS_CNFG.RAW_MAX : Raw maximum value from AI card
   // RIO_03.FIRST_TANK.DECK_IG_PRESS_CNFG.NORM : Normalised real value
   // RIO_03.FIRST_TANK.DECK_IG_PRESS_CNFG.ENG_MIN : Engineering units minimum value
   // RIO_03.FIRST_TANK.DECK_IG_PRESS_CNFG.ENG_MAX : Engineering units maximum value
   // RIO_03.FIRST_TANK.TANKS_PRESS_CNFG : Tank Group Pressure (PT-424)
   // RIO_03.FIRST_TANK.TANKS_PRESS_CNFG.RAW_MIN : Raw minimum value from AI card
   // RIO_03.FIRST_TANK.TANKS_PRESS_CNFG.RAW_MAX : Raw maximum value from AI card
   // RIO_03.FIRST_TANK.TANKS_PRESS_CNFG.NORM : Normalised real value
   // RIO_03.FIRST_TANK.TANKS_PRESS_CNFG.ENG_MIN : Engineering units minimum value
   // RIO_03.FIRST_TANK.TANKS_PRESS_CNFG.ENG_MAX : Engineering units maximum value
   // RIO_04.FIRST_TANK.O2_MONITOR : Space monitor, 600-Tx-433
   // RIO_04.FIRST_TANK.DECK_IG_PRESS : Deck main IG pressure, PT-415
   // RIO_04.FIRST_TANK.TANKS_PRESS : Tank group pressure, PT-424
   // RIO_04.FIRST_TANK.TANKS_PRESS_HIHI : Tank group pressure, PS-436
   // RIO_04.FIRST_TANK.TANK_GROUP_SPARE_DI_2 : Spare input
   // RIO_04.FIRST_TANK.TANK_GROUP_SPARE_DI_3 : Spare input
   // RIO_04.FIRST_TANK.TANK_GROUP_SPARE_DI_4 : Spare input
   // RIO_04.FIRST_TANK.TANK_GROUP_SPARE_DI_5 : Spare input
   // RIO_04.FIRST_TANK.TANK_GROUP_SPARE_DI_6 : Spare input
   // RIO_04.FIRST_TANK.TANK_GROUP_SPARE_DI_7 : Spare input
   // RIO_04.FIRST_TANK.GTT_ISOL_VALVE_OPEN : Gas to tank isolation valve feedback, CV-422
   // RIO_04.FIRST_TANK.GTT_ISOL_VALVE_CLSD : Gas to tank isolation valve feedback, CV-422
   // RIO_04.FIRST_TANK.TANK_VENT_A_OPEN : Tank vent valve feedback, CV-441-A
   // RIO_04.FIRST_TANK.TANK_VENT_A_CLSD : Tank vent valve feedback, CV-441-A
   // RIO_04.FIRST_TANK.TANK_VENT_B_OPEN : Tank vent valve feedback, CV-441-B
   // RIO_04.FIRST_TANK.TANK_VENT_B_CLSD : Tank vent valve feedback, CV-441-B
   // RIO_04.FIRST_TANK.BWT_LEVEL_HIHI : Tank water level, LS-425
   // RIO_04.FIRST_TANK.TANK_ALARM : Spare input
   // RIO_04.FIRST_TANK.SPARE_DI_7 : Spare input
   // RIO_04.FIRST_TANK.USD_FLOW : FIT-418
   // RIO_04.FIRST_TANK.MBG_FLOW : FIT-420